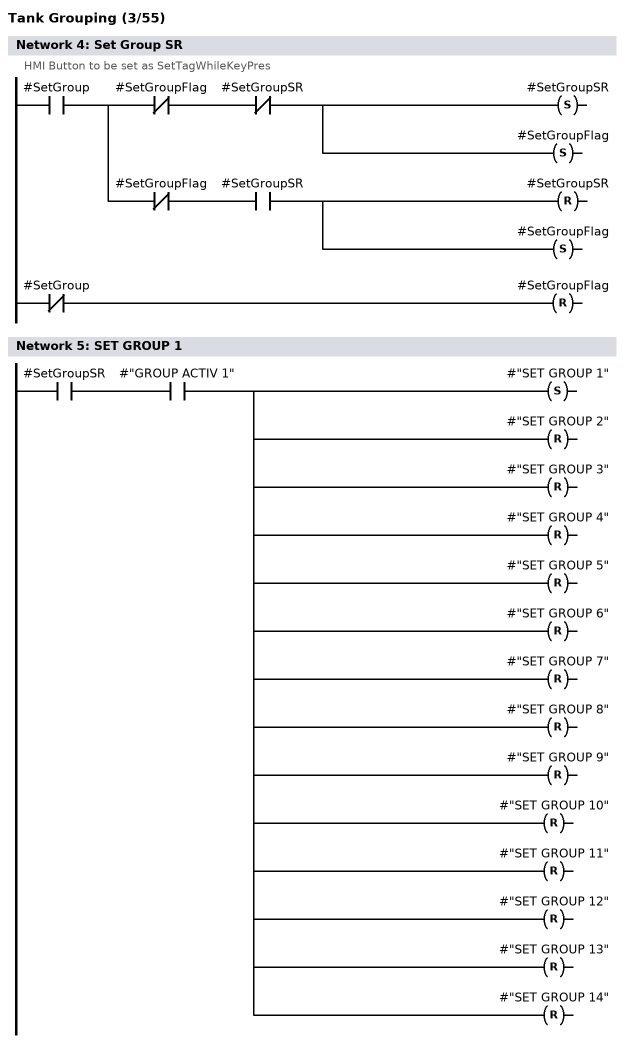
   RUNG wire#powerrail
      Contact( #SetGroup )
      wire#w1
      I_Contact( #SetGroupFlag )
      I_Contact( #SetGroupSR )
      wire#w2
      S_Coil( #SetGroupSR )
   END_RUNG
   RUNG wire#w2
      S_Coil( #SetGroupFlag )
   END_RUNG
   RUNG wire#w1
      I_Contact( #SetGroupFlag )
      Contact( #SetGroupSR )
      wire#w3
      R_Coil( #SetGroupSR )
   END_RUNG
   RUNG wire#w3
      S_Coil( #SetGroupFlag )
   END_RUNG
   RUNG wire#powerrail
      I_Contact( #SetGroup )
      R_Coil( #SetGroupFlag )
   END_RUNG
   // the same network as SCL:
   #_w1 := #SetGroup AND NOT #SetGroupFlag AND NOT #SetGroupSR;
   IF #_w1 THEN
       #SetGroupSR := TRUE;
       #SetGroupFlag := TRUE;
   END_IF;
   #_w2 := #SetGroup AND NOT #SetGroupFlag AND #SetGroupSR;
   IF #_w2 THEN
       #SetGroupSR := FALSE;
       #SetGroupFlag := TRUE;
   END_IF;
   IF NOT #SetGroup THEN #SetGroupFlag := FALSE; END_IF;
END_REGION

REGION Network 5: SET GROUP 1
   RUNG wire#powerrail
      Contact( #SetGroupSR )
      Contact( #"GROUP ACTIV 1" )
      wire#w1
      S_Coil( #"SET GROUP 1" )
   END_RUNG
   RUNG wire#w1
      R_Coil( #"SET GROUP 2" )
   END_RUNG
   RUNG wire#w1
      R_Coil( #"SET GROUP 3" )
   END_RUNG
   RUNG wire#w1
      R_Coil( #"SET GROUP 4" )
   END_RUNG
   RUNG wire#w1
      R_Coil( #"SET GROUP 5" )
   END_RUNG
   RUNG wire#w1
      R_Coil( #"SET GROUP 6" )
   END_RUNG
   RUNG wire#w1
      R_Coil( #"SET GROUP 7" )
   END_RUNG
   RUNG wire#w1
      R_Coil( #"SET GROUP 8" )
   END_RUNG
   RUNG wire#w1
      R_Coil( #"SET GROUP 9" )
   END_RUNG
   RUNG wire#w1
      R_Coil( #"SET GROUP 10" )
   END_RUNG
   RUNG wire#w1
      R_Coil( #"SET GROUP 11" )
   END_RUNG
   RUNG wire#w1
      R_Coil( #"SET GROUP 12" )
   END_RUNG
   RUNG wire#w1
      R_Coil( #"SET GROUP 13" )
   END_RUNG
   RUNG wire#w1
      R_Coil( #"SET GROUP 14" )
   END_RUNG
   // the same network as SCL:
   IF #SetGroupSR AND #"GROUP ACTIV 1" THEN
       #"SET GROUP 1" := TRUE;
       #"SET GROUP 2" := FALSE;
       #"SET GROUP 3" := FALSE;
       #"SET GROUP 4" := FALSE;
       #"SET GROUP 5" := FALSE;
       #"SET GROUP 6" := FALSE;
       #"SET GROUP 7" := FALSE;
       #"SET GROUP 8" := FALSE;
       #"SET GROUP 9" := FALSE;
       #"SET GROUP 10" := FALSE;
       #"SET GROUP 11" := FALSE;
       #"SET GROUP 12" := FALSE;
       #"SET GROUP 13" := FALSE;
       #"SET GROUP 14" := FALSE;
   END_IF;
END_REGION

REGION Network 6: SET GROUP 2
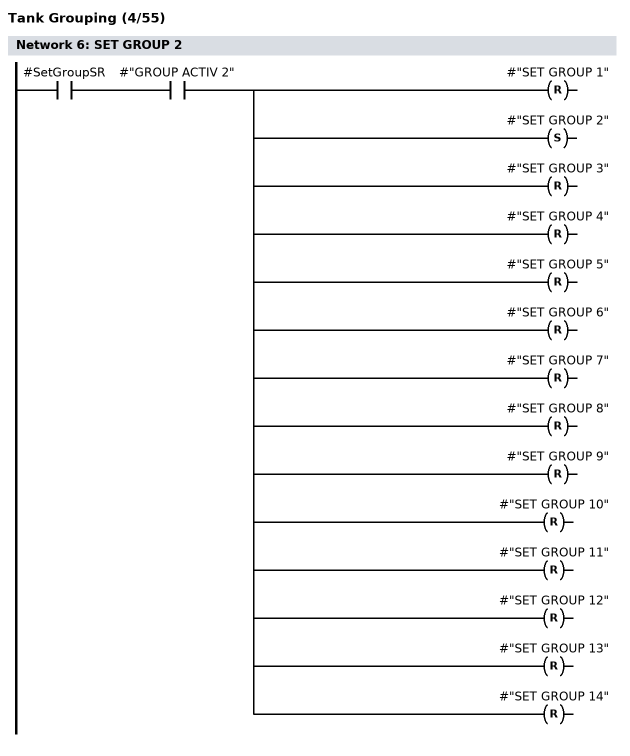
   RUNG wire#powerrail
      Contact( #SetGroupSR )
      Contact( #"GROUP ACTIV 2" )
      wire#w1
      R_Coil( #"SET GROUP 1" )
   END_RUNG
   RUNG wire#w1
      S_Coil( #"SET GROUP 2" )
   END_RUNG
   RUNG wire#w1
      R_Coil( #"SET GROUP 3" )
   END_RUNG
   RUNG wire#w1
      R_Coil( #"SET GROUP 4" )
   END_RUNG
   RUNG wire#w1
      R_Coil( #"SET GROUP 5" )
   END_RUNG
   RUNG wire#w1
      R_Coil( #"SET GROUP 6" )
   END_RUNG
   RUNG wire#w1
      R_Coil( #"SET GROUP 7" )
   END_RUNG
   RUNG wire#w1
      R_Coil( #"SET GROUP 8" )
   END_RUNG
   RUNG wire#w1
      R_Coil( #"SET GROUP 9" )
   END_RUNG
   RUNG wire#w1
      R_Coil( #"SET GROUP 10" )
   END_RUNG
   RUNG wire#w1
      R_Coil( #"SET GROUP 11" )
   END_RUNG
   RUNG wire#w1
      R_Coil( #"SET GROUP 12" )
   END_RUNG
   RUNG wire#w1
      R_Coil( #"SET GROUP 13" )
   END_RUNG
   RUNG wire#w1
      R_Coil( #"SET GROUP 14" )
   END_RUNG
   // the same network as SCL:
   IF #SetGroupSR AND #"GROUP ACTIV 2" THEN
       #"SET GROUP 1" := FALSE;
       #"SET GROUP 2" := TRUE;
       #"SET GROUP 3" := FALSE;
       #"SET GROUP 4" := FALSE;
       #"SET GROUP 5" := FALSE;
       #"SET GROUP 6" := FALSE;
       #"SET GROUP 7" := FALSE;
       #"SET GROUP 8" := FALSE;
       #"SET GROUP 9" := FALSE;
       #"SET GROUP 10" := FALSE;
       #"SET GROUP 11" := FALSE;
       #"SET GROUP 12" := FALSE;
       #"SET GROUP 13" := FALSE;
       #"SET GROUP 14" := FALSE;
   END_IF;
END_REGION

REGION Network 7: SET GROUP 3
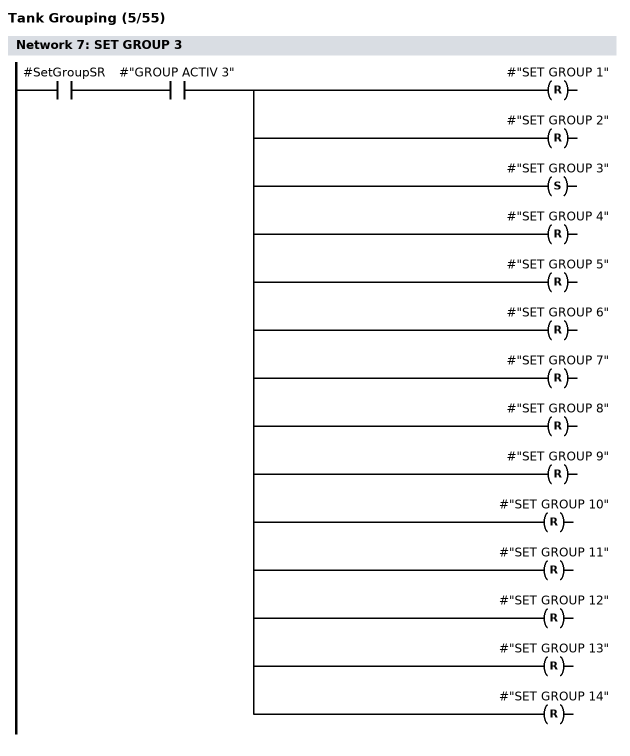
   RUNG wire#powerrail
      Contact( #SetGroupSR )
      Contact( #"GROUP ACTIV 3" )
      wire#w1
      R_Coil( #"SET GROUP 1" )
   END_RUNG
   RUNG wire#w1
      R_Coil( #"SET GROUP 2" )
   END_RUNG
   RUNG wire#w1
      S_Coil( #"SET GROUP 3" )
   END_RUNG
   RUNG wire#w1
      R_Coil( #"SET GROUP 4" )
   END_RUNG
   RUNG wire#w1
      R_Coil( #"SET GROUP 5" )
   END_RUNG
   RUNG wire#w1
      R_Coil( #"SET GROUP 6" )
   END_RUNG
   RUNG wire#w1
      R_Coil( #"SET GROUP 7" )
   END_RUNG
   RUNG wire#w1
      R_Coil( #"SET GROUP 8" )
   END_RUNG
   RUNG wire#w1
      R_Coil( #"SET GROUP 9" )
   END_RUNG
   RUNG wire#w1
      R_Coil( #"SET GROUP 10" )
   END_RUNG
   RUNG wire#w1
      R_Coil( #"SET GROUP 11" )
   END_RUNG
   RUNG wire#w1
      R_Coil( #"SET GROUP 12" )
   END_RUNG
   RUNG wire#w1
      R_Coil( #"SET GROUP 13" )
   END_RUNG
   RUNG wire#w1
      R_Coil( #"SET GROUP 14" )
   END_RUNG
   // the same network as SCL:
   IF #SetGroupSR AND #"GROUP ACTIV 3" THEN
       #"SET GROUP 1" := FALSE;
       #"SET GROUP 2" := FALSE;
       #"SET GROUP 3" := TRUE;
       #"SET GROUP 4" := FALSE;
       #"SET GROUP 5" := FALSE;
       #"SET GROUP 6" := FALSE;
       #"SET GROUP 7" := FALSE;
       #"SET GROUP 8" := FALSE;
       #"SET GROUP 9" := FALSE;
       #"SET GROUP 10" := FALSE;
       #"SET GROUP 11" := FALSE;
       #"SET GROUP 12" := FALSE;
       #"SET GROUP 13" := FALSE;
       #"SET GROUP 14" := FALSE;
   END_IF;
END_REGION

REGION Network 8: SET GROUP 4
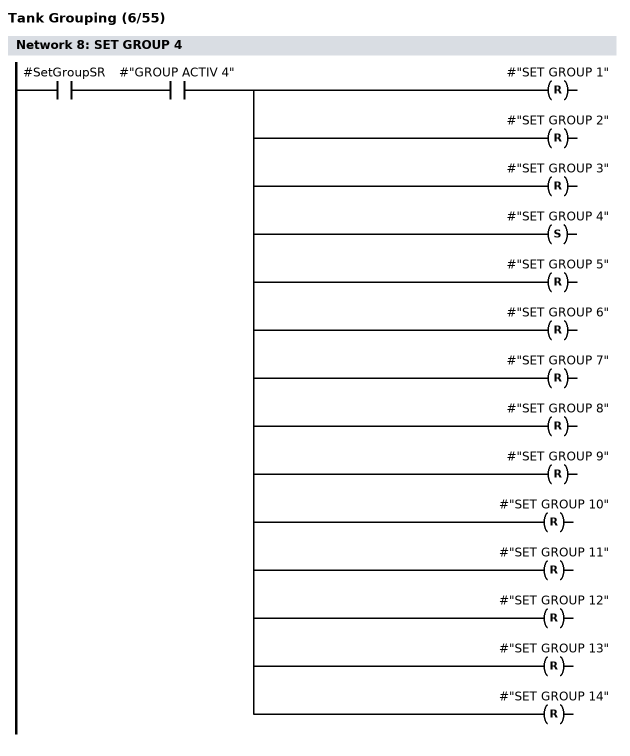
   RUNG wire#powerrail
      Contact( #SetGroupSR )
      Contact( #"GROUP ACTIV 4" )
      wire#w1
      R_Coil( #"SET GROUP 1" )
   END_RUNG
   RUNG wire#w1
      R_Coil( #"SET GROUP 2" )
   END_RUNG
   RUNG wire#w1
      R_Coil( #"SET GROUP 3" )
   END_RUNG
   RUNG wire#w1
      S_Coil( #"SET GROUP 4" )
   END_RUNG
   RUNG wire#w1
      R_Coil( #"SET GROUP 5" )
   END_RUNG
   RUNG wire#w1
      R_Coil( #"SET GROUP 6" )
   END_RUNG
   RUNG wire#w1
      R_Coil( #"SET GROUP 7" )
   END_RUNG
   RUNG wire#w1
      R_Coil( #"SET GROUP 8" )
   END_RUNG
   RUNG wire#w1
      R_Coil( #"SET GROUP 9" )
   END_RUNG
   RUNG wire#w1
      R_Coil( #"SET GROUP 10" )
   END_RUNG
   RUNG wire#w1
      R_Coil( #"SET GROUP 11" )
   END_RUNG
   RUNG wire#w1
      R_Coil( #"SET GROUP 12" )
   END_RUNG
   RUNG wire#w1
      R_Coil( #"SET GROUP 13" )
   END_RUNG
   RUNG wire#w1
      R_Coil( #"SET GROUP 14" )
   END_RUNG
   // the same network as SCL:
   IF #SetGroupSR AND #"GROUP ACTIV 4" THEN
       #"SET GROUP 1" := FALSE;
       #"SET GROUP 2" := FALSE;
       #"SET GROUP 3" := FALSE;
       #"SET GROUP 4" := TRUE;
       #"SET GROUP 5" := FALSE;
       #"SET GROUP 6" := FALSE;
       #"SET GROUP 7" := FALSE;
       #"SET GROUP 8" := FALSE;
       #"SET GROUP 9" := FALSE;
       #"SET GROUP 10" := FALSE;
       #"SET GROUP 11" := FALSE;
       #"SET GROUP 12" := FALSE;
       #"SET GROUP 13" := FALSE;
       #"SET GROUP 14" := FALSE;
   END_IF;
END_REGION

REGION Network 9: SET GROUP 5
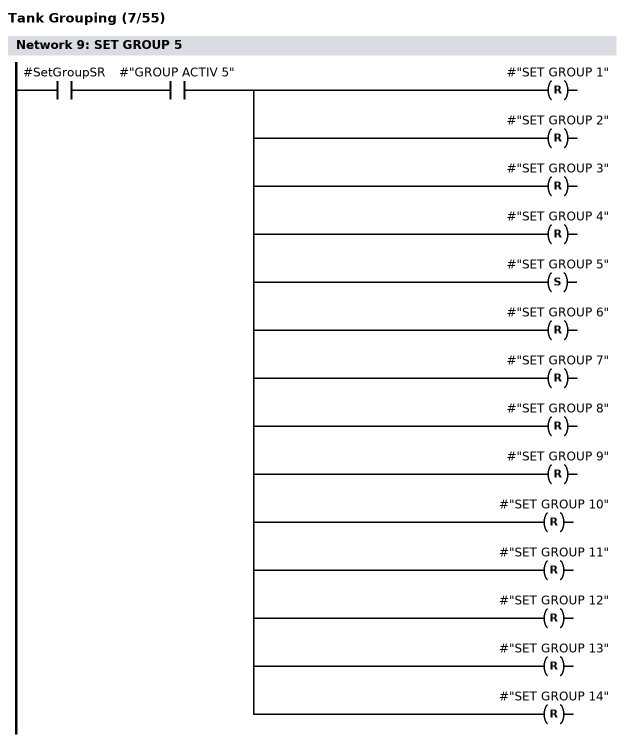
   RUNG wire#powerrail
      Contact( #SetGroupSR )
      Contact( #"GROUP ACTIV 5" )
      wire#w1
      R_Coil( #"SET GROUP 1" )
   END_RUNG
   RUNG wire#w1
      R_Coil( #"SET GROUP 2" )
   END_RUNG
   RUNG wire#w1
      R_Coil( #"SET GROUP 3" )
   END_RUNG
   RUNG wire#w1
      R_Coil( #"SET GROUP 4" )
   END_RUNG
   RUNG wire#w1
      S_Coil( #"SET GROUP 5" )
   END_RUNG
   RUNG wire#w1
      R_Coil( #"SET GROUP 6" )
   END_RUNG
   RUNG wire#w1
      R_Coil( #"SET GROUP 7" )
   END_RUNG
   RUNG wire#w1
      R_Coil( #"SET GROUP 8" )
   END_RUNG
   RUNG wire#w1
      R_Coil( #"SET GROUP 9" )
   END_RUNG
   RUNG wire#w1
      R_Coil( #"SET GROUP 10" )
   END_RUNG
   RUNG wire#w1
      R_Coil( #"SET GROUP 11" )
   END_RUNG
   RUNG wire#w1
      R_Coil( #"SET GROUP 12" )
   END_RUNG
   RUNG wire#w1
      R_Coil( #"SET GROUP 13" )
   END_RUNG
   RUNG wire#w1
      R_Coil( #"SET GROUP 14" )
   END_RUNG
   // the same network as SCL:
   IF #SetGroupSR AND #"GROUP ACTIV 5" THEN
       #"SET GROUP 1" := FALSE;
       #"SET GROUP 2" := FALSE;
       #"SET GROUP 3" := FALSE;
       #"SET GROUP 4" := FALSE;
       #"SET GROUP 5" := TRUE;
       #"SET GROUP 6" := FALSE;
       #"SET GROUP 7" := FALSE;
       #"SET GROUP 8" := FALSE;
       #"SET GROUP 9" := FALSE;
       #"SET GROUP 10" := FALSE;
       #"SET GROUP 11" := FALSE;
       #"SET GROUP 12" := FALSE;
       #"SET GROUP 13" := FALSE;
       #"SET GROUP 14" := FALSE;
   END_IF;
END_REGION

REGION Network 10: SET GROUP 6
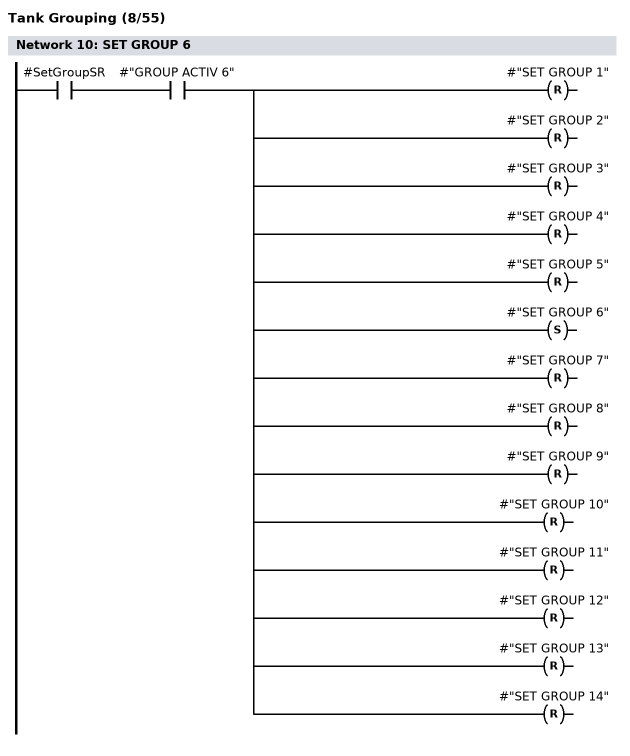
   RUNG wire#powerrail
      Contact( #SetGroupSR )
      Contact( #"GROUP ACTIV 6" )
      wire#w1
      R_Coil( #"SET GROUP 1" )
   END_RUNG
   RUNG wire#w1
      R_Coil( #"SET GROUP 2" )
   END_RUNG
   RUNG wire#w1
      R_Coil( #"SET GROUP 3" )
   END_RUNG
   RUNG wire#w1
      R_Coil( #"SET GROUP 4" )
   END_RUNG
   RUNG wire#w1
      R_Coil( #"SET GROUP 5" )
   END_RUNG
   RUNG wire#w1
      S_Coil( #"SET GROUP 6" )
   END_RUNG
   RUNG wire#w1
      R_Coil( #"SET GROUP 7" )
   END_RUNG
   RUNG wire#w1
      R_Coil( #"SET GROUP 8" )
   END_RUNG
   RUNG wire#w1
      R_Coil( #"SET GROUP 9" )
   END_RUNG
   RUNG wire#w1
      R_Coil( #"SET GROUP 10" )
   END_RUNG
   RUNG wire#w1
      R_Coil( #"SET GROUP 11" )
   END_RUNG
   RUNG wire#w1
      R_Coil( #"SET GROUP 12" )
   END_RUNG
   RUNG wire#w1
      R_Coil( #"SET GROUP 13" )
   END_RUNG
   RUNG wire#w1
      R_Coil( #"SET GROUP 14" )
   END_RUNG
   // the same network as SCL:
   IF #SetGroupSR AND #"GROUP ACTIV 6" THEN
       #"SET GROUP 1" := FALSE;
       #"SET GROUP 2" := FALSE;
       #"SET GROUP 3" := FALSE;
       #"SET GROUP 4" := FALSE;
       #"SET GROUP 5" := FALSE;
       #"SET GROUP 6" := TRUE;
       #"SET GROUP 7" := FALSE;
       #"SET GROUP 8" := FALSE;
       #"SET GROUP 9" := FALSE;
       #"SET GROUP 10" := FALSE;
       #"SET GROUP 11" := FALSE;
       #"SET GROUP 12" := FALSE;
       #"SET GROUP 13" := FALSE;
       #"SET GROUP 14" := FALSE;
   END_IF;
END_REGION

REGION Network 11: SET GROUP 7
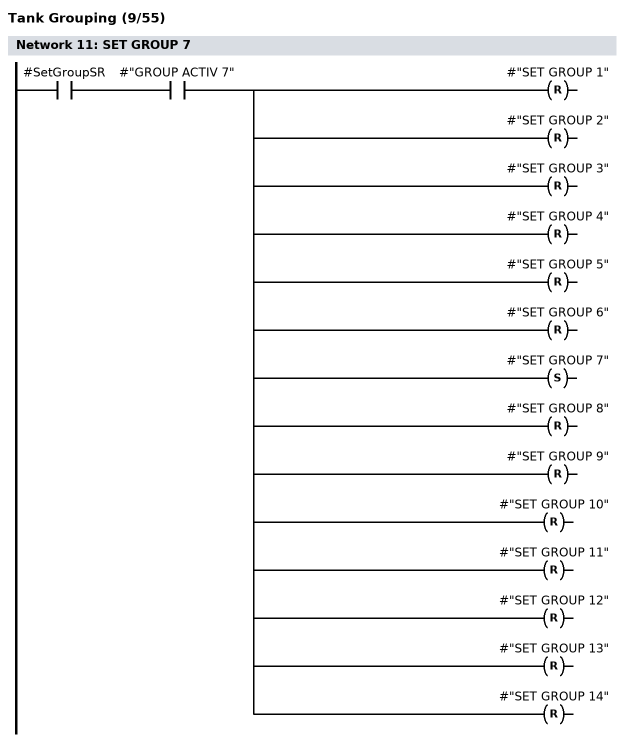
   RUNG wire#powerrail
      Contact( #SetGroupSR )
      Contact( #"GROUP ACTIV 7" )
      wire#w1
      R_Coil( #"SET GROUP 1" )
   END_RUNG
   RUNG wire#w1
      R_Coil( #"SET GROUP 2" )
   END_RUNG
   RUNG wire#w1
      R_Coil( #"SET GROUP 3" )
   END_RUNG
   RUNG wire#w1
      R_Coil( #"SET GROUP 4" )
   END_RUNG
   RUNG wire#w1
      R_Coil( #"SET GROUP 5" )
   END_RUNG
   RUNG wire#w1
      R_Coil( #"SET GROUP 6" )
   END_RUNG
   RUNG wire#w1
      S_Coil( #"SET GROUP 7" )
   END_RUNG
   RUNG wire#w1
      R_Coil( #"SET GROUP 8" )
   END_RUNG
   RUNG wire#w1
      R_Coil( #"SET GROUP 9" )
   END_RUNG
   RUNG wire#w1
      R_Coil( #"SET GROUP 10" )
   END_RUNG
   RUNG wire#w1
      R_Coil( #"SET GROUP 11" )
   END_RUNG
   RUNG wire#w1
      R_Coil( #"SET GROUP 12" )
   END_RUNG
   RUNG wire#w1
      R_Coil( #"SET GROUP 13" )
   END_RUNG
   RUNG wire#w1
      R_Coil( #"SET GROUP 14" )
   END_RUNG
   // the same network as SCL:
   IF #SetGroupSR AND #"GROUP ACTIV 7" THEN
       #"SET GROUP 1" := FALSE;
       #"SET GROUP 2" := FALSE;
       #"SET GROUP 3" := FALSE;
       #"SET GROUP 4" := FALSE;
       #"SET GROUP 5" := FALSE;
       #"SET GROUP 6" := FALSE;
       #"SET GROUP 7" := TRUE;
       #"SET GROUP 8" := FALSE;
       #"SET GROUP 9" := FALSE;
       #"SET GROUP 10" := FALSE;
       #"SET GROUP 11" := FALSE;
       #"SET GROUP 12" := FALSE;
       #"SET GROUP 13" := FALSE;
       #"SET GROUP 14" := FALSE;
   END_IF;
END_REGION

REGION Network 12: SET GROUP 8
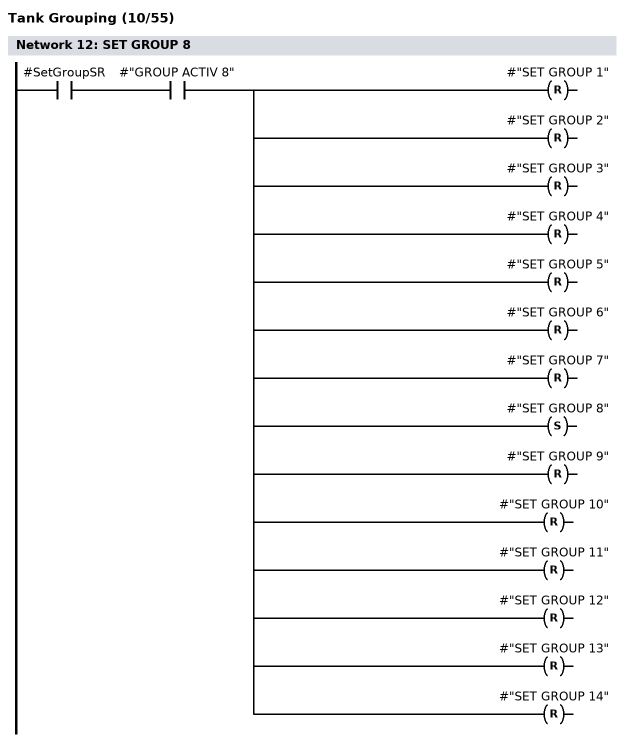
   RUNG wire#powerrail
      Contact( #SetGroupSR )
      Contact( #"GROUP ACTIV 8" )
      wire#w1
      R_Coil( #"SET GROUP 1" )
   END_RUNG
   RUNG wire#w1
      R_Coil( #"SET GROUP 2" )
   END_RUNG
   RUNG wire#w1
      R_Coil( #"SET GROUP 3" )
   END_RUNG
   RUNG wire#w1
      R_Coil( #"SET GROUP 4" )
   END_RUNG
   RUNG wire#w1
      R_Coil( #"SET GROUP 5" )
   END_RUNG
   RUNG wire#w1
      R_Coil( #"SET GROUP 6" )
   END_RUNG
   RUNG wire#w1
      R_Coil( #"SET GROUP 7" )
   END_RUNG
   RUNG wire#w1
      S_Coil( #"SET GROUP 8" )
   END_RUNG
   RUNG wire#w1
      R_Coil( #"SET GROUP 9" )
   END_RUNG
   RUNG wire#w1
      R_Coil( #"SET GROUP 10" )
   END_RUNG
   RUNG wire#w1
      R_Coil( #"SET GROUP 11" )
   END_RUNG
   RUNG wire#w1
      R_Coil( #"SET GROUP 12" )
   END_RUNG
   RUNG wire#w1
      R_Coil( #"SET GROUP 13" )
   END_RUNG
   RUNG wire#w1
      R_Coil( #"SET GROUP 14" )
   END_RUNG
   // the same network as SCL:
   IF #SetGroupSR AND #"GROUP ACTIV 8" THEN
       #"SET GROUP 1" := FALSE;
       #"SET GROUP 2" := FALSE;
       #"SET GROUP 3" := FALSE;
       #"SET GROUP 4" := FALSE;
       #"SET GROUP 5" := FALSE;
       #"SET GROUP 6" := FALSE;
       #"SET GROUP 7" := FALSE;
       #"SET GROUP 8" := TRUE;
       #"SET GROUP 9" := FALSE;
       #"SET GROUP 10" := FALSE;
       #"SET GROUP 11" := FALSE;
       #"SET GROUP 12" := FALSE;
       #"SET GROUP 13" := FALSE;
       #"SET GROUP 14" := FALSE;
   END_IF;
END_REGION

REGION Network 13: SET GROUP 9
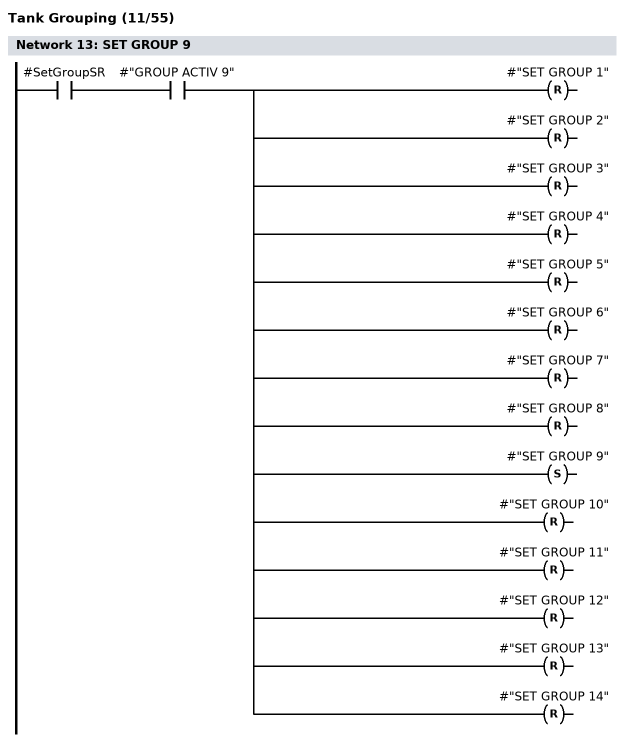
   RUNG wire#powerrail
      Contact( #SetGroupSR )
      Contact( #"GROUP ACTIV 9" )
      wire#w1
      R_Coil( #"SET GROUP 1" )
   END_RUNG
   RUNG wire#w1
      R_Coil( #"SET GROUP 2" )
   END_RUNG
   RUNG wire#w1
      R_Coil( #"SET GROUP 3" )
   END_RUNG
   RUNG wire#w1
      R_Coil( #"SET GROUP 4" )
   END_RUNG
   RUNG wire#w1
      R_Coil( #"SET GROUP 5" )
   END_RUNG
   RUNG wire#w1
      R_Coil( #"SET GROUP 6" )
   END_RUNG
   RUNG wire#w1
      R_Coil( #"SET GROUP 7" )
   END_RUNG
   RUNG wire#w1
      R_Coil( #"SET GROUP 8" )
   END_RUNG
   RUNG wire#w1
      S_Coil( #"SET GROUP 9" )
   END_RUNG
   RUNG wire#w1
      R_Coil( #"SET GROUP 10" )
   END_RUNG
   RUNG wire#w1
      R_Coil( #"SET GROUP 11" )
   END_RUNG
   RUNG wire#w1
      R_Coil( #"SET GROUP 12" )
   END_RUNG
   RUNG wire#w1
      R_Coil( #"SET GROUP 13" )
   END_RUNG
   RUNG wire#w1
      R_Coil( #"SET GROUP 14" )
   END_RUNG
   // the same network as SCL:
   IF #SetGroupSR AND #"GROUP ACTIV 9" THEN
       #"SET GROUP 1" := FALSE;
       #"SET GROUP 2" := FALSE;
       #"SET GROUP 3" := FALSE;
       #"SET GROUP 4" := FALSE;
       #"SET GROUP 5" := FALSE;
       #"SET GROUP 6" := FALSE;
       #"SET GROUP 7" := FALSE;
       #"SET GROUP 8" := FALSE;
       #"SET GROUP 9" := TRUE;
       #"SET GROUP 10" := FALSE;
       #"SET GROUP 11" := FALSE;
       #"SET GROUP 12" := FALSE;
       #"SET GROUP 13" := FALSE;
       #"SET GROUP 14" := FALSE;
   END_IF;
END_REGION

REGION Network 14: SET GROUP 10
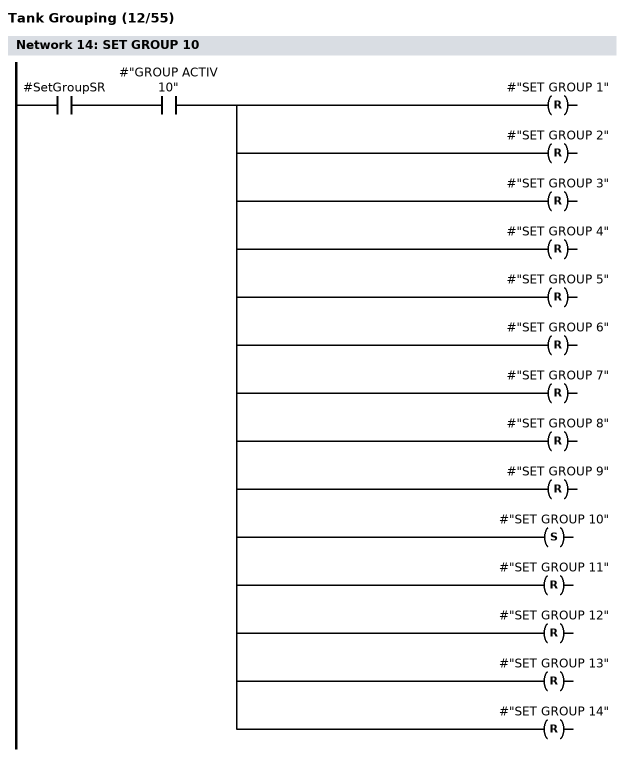
   RUNG wire#powerrail
      Contact( #SetGroupSR )
      Contact( #"GROUP ACTIV 10" )
      wire#w1
      R_Coil( #"SET GROUP 1" )
   END_RUNG
   RUNG wire#w1
      R_Coil( #"SET GROUP 2" )
   END_RUNG
   RUNG wire#w1
      R_Coil( #"SET GROUP 3" )
   END_RUNG
   RUNG wire#w1
      R_Coil( #"SET GROUP 4" )
   END_RUNG
   RUNG wire#w1
      R_Coil( #"SET GROUP 5" )
   END_RUNG
   RUNG wire#w1
      R_Coil( #"SET GROUP 6" )
   END_RUNG
   RUNG wire#w1
      R_Coil( #"SET GROUP 7" )
   END_RUNG
   RUNG wire#w1
      R_Coil( #"SET GROUP 8" )
   END_RUNG
   RUNG wire#w1
      R_Coil( #"SET GROUP 9" )
   END_RUNG
   RUNG wire#w1
      S_Coil( #"SET GROUP 10" )
   END_RUNG
   RUNG wire#w1
      R_Coil( #"SET GROUP 11" )
   END_RUNG
   RUNG wire#w1
      R_Coil( #"SET GROUP 12" )
   END_RUNG
   RUNG wire#w1
      R_Coil( #"SET GROUP 13" )
   END_RUNG
   RUNG wire#w1
      R_Coil( #"SET GROUP 14" )
   END_RUNG
   // the same network as SCL:
   IF #SetGroupSR AND #"GROUP ACTIV 10" THEN
       #"SET GROUP 1" := FALSE;
       #"SET GROUP 2" := FALSE;
       #"SET GROUP 3" := FALSE;
       #"SET GROUP 4" := FALSE;
       #"SET GROUP 5" := FALSE;
       #"SET GROUP 6" := FALSE;
       #"SET GROUP 7" := FALSE;
       #"SET GROUP 8" := FALSE;
       #"SET GROUP 9" := FALSE;
       #"SET GROUP 10" := TRUE;
       #"SET GROUP 11" := FALSE;
       #"SET GROUP 12" := FALSE;
       #"SET GROUP 13" := FALSE;
       #"SET GROUP 14" := FALSE;
   END_IF;
END_REGION

REGION Network 15: SET GROUP 11
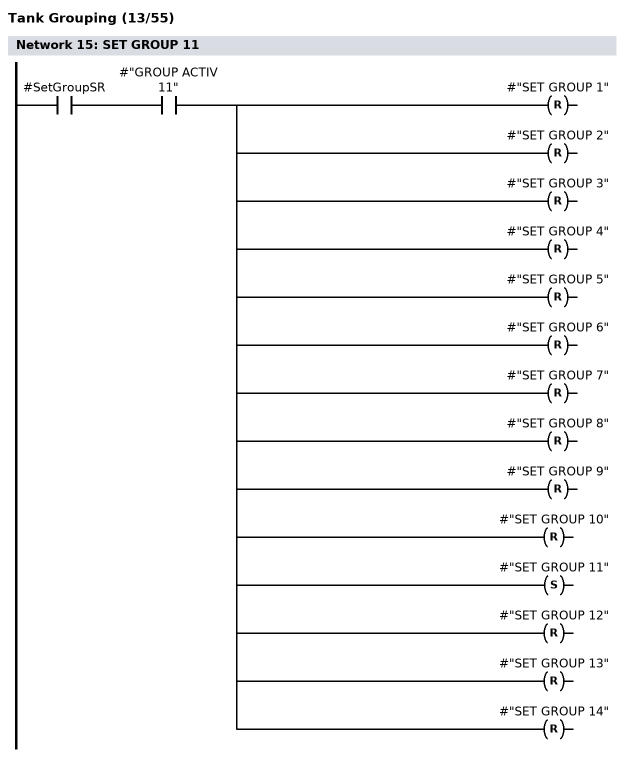
   RUNG wire#powerrail
      Contact( #SetGroupSR )
      Contact( #"GROUP ACTIV 11" )
      wire#w1
      R_Coil( #"SET GROUP 1" )
   END_RUNG
   RUNG wire#w1
      R_Coil( #"SET GROUP 2" )
   END_RUNG
   RUNG wire#w1
      R_Coil( #"SET GROUP 3" )
   END_RUNG
   RUNG wire#w1
      R_Coil( #"SET GROUP 4" )
   END_RUNG
   RUNG wire#w1
      R_Coil( #"SET GROUP 5" )
   END_RUNG
   RUNG wire#w1
      R_Coil( #"SET GROUP 6" )
   END_RUNG
   RUNG wire#w1
      R_Coil( #"SET GROUP 7" )
   END_RUNG
   RUNG wire#w1
      R_Coil( #"SET GROUP 8" )
   END_RUNG
   RUNG wire#w1
      R_Coil( #"SET GROUP 9" )
   END_RUNG
   RUNG wire#w1
      R_Coil( #"SET GROUP 10" )
   END_RUNG
   RUNG wire#w1
      S_Coil( #"SET GROUP 11" )
   END_RUNG
   RUNG wire#w1
      R_Coil( #"SET GROUP 12" )
   END_RUNG
   RUNG wire#w1
      R_Coil( #"SET GROUP 13" )
   END_RUNG
   RUNG wire#w1
      R_Coil( #"SET GROUP 14" )
   END_RUNG
   // the same network as SCL:
   IF #SetGroupSR AND #"GROUP ACTIV 11" THEN
       #"SET GROUP 1" := FALSE;
       #"SET GROUP 2" := FALSE;
       #"SET GROUP 3" := FALSE;
       #"SET GROUP 4" := FALSE;
       #"SET GROUP 5" := FALSE;
       #"SET GROUP 6" := FALSE;
       #"SET GROUP 7" := FALSE;
       #"SET GROUP 8" := FALSE;
       #"SET GROUP 9" := FALSE;
       #"SET GROUP 10" := FALSE;
       #"SET GROUP 11" := TRUE;
       #"SET GROUP 12" := FALSE;
       #"SET GROUP 13" := FALSE;
       #"SET GROUP 14" := FALSE;
   END_IF;
END_REGION

REGION Network 16: SET GROUP 12
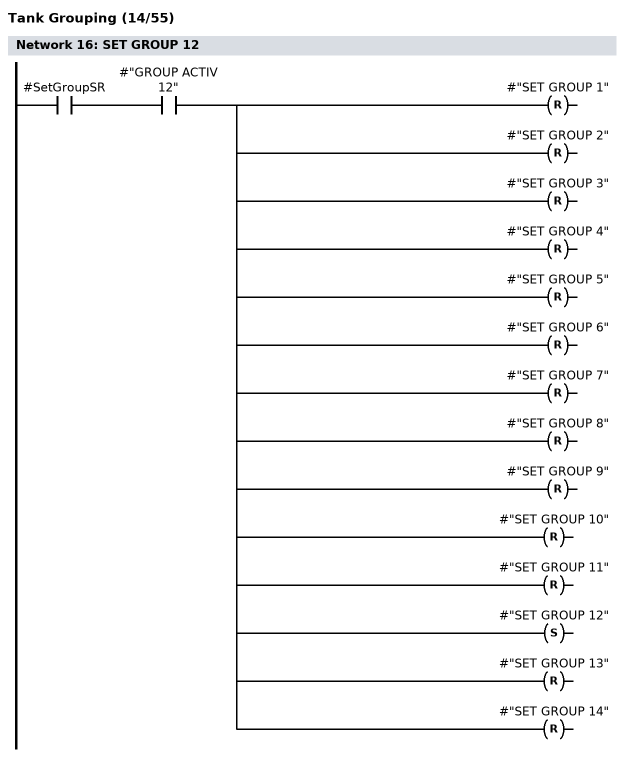
   RUNG wire#powerrail
      Contact( #SetGroupSR )
      Contact( #"GROUP ACTIV 12" )
      wire#w1
      R_Coil( #"SET GROUP 1" )
   END_RUNG
   RUNG wire#w1
      R_Coil( #"SET GROUP 2" )
   END_RUNG
   RUNG wire#w1
      R_Coil( #"SET GROUP 3" )
   END_RUNG
   RUNG wire#w1
      R_Coil( #"SET GROUP 4" )
   END_RUNG
   RUNG wire#w1
      R_Coil( #"SET GROUP 5" )
   END_RUNG
   RUNG wire#w1
      R_Coil( #"SET GROUP 6" )
   END_RUNG
   RUNG wire#w1
      R_Coil( #"SET GROUP 7" )
   END_RUNG
   RUNG wire#w1
      R_Coil( #"SET GROUP 8" )
   END_RUNG
   RUNG wire#w1
      R_Coil( #"SET GROUP 9" )
   END_RUNG
   RUNG wire#w1
      R_Coil( #"SET GROUP 10" )
   END_RUNG
   RUNG wire#w1
      R_Coil( #"SET GROUP 11" )
   END_RUNG
   RUNG wire#w1
      S_Coil( #"SET GROUP 12" )
   END_RUNG
   RUNG wire#w1
      R_Coil( #"SET GROUP 13" )
   END_RUNG
   RUNG wire#w1
      R_Coil( #"SET GROUP 14" )
   END_RUNG
   // the same network as SCL:
   IF #SetGroupSR AND #"GROUP ACTIV 12" THEN
       #"SET GROUP 1" := FALSE;
       #"SET GROUP 2" := FALSE;
       #"SET GROUP 3" := FALSE;
       #"SET GROUP 4" := FALSE;
       #"SET GROUP 5" := FALSE;
       #"SET GROUP 6" := FALSE;
       #"SET GROUP 7" := FALSE;
       #"SET GROUP 8" := FALSE;
       #"SET GROUP 9" := FALSE;
       #"SET GROUP 10" := FALSE;
       #"SET GROUP 11" := FALSE;
       #"SET GROUP 12" := TRUE;
       #"SET GROUP 13" := FALSE;
       #"SET GROUP 14" := FALSE;
   END_IF;
END_REGION

REGION Network 17: SET GROUP 13
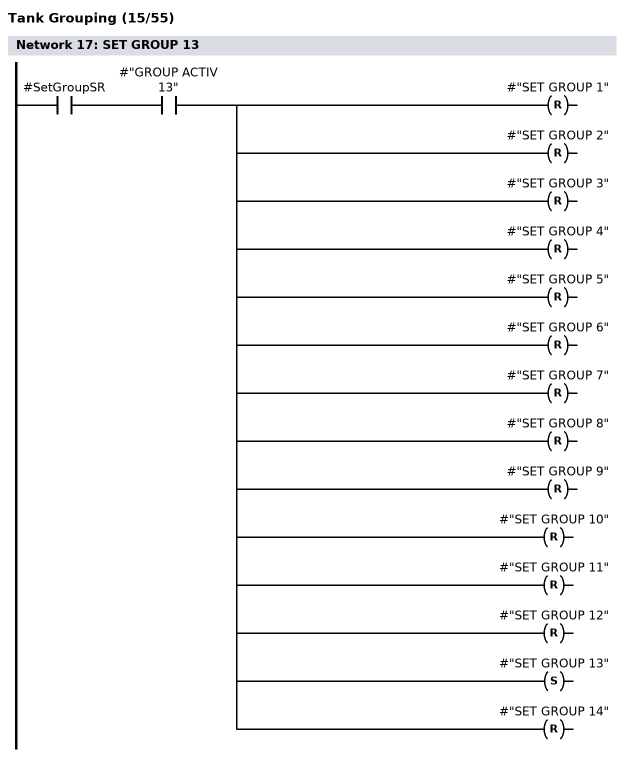
   RUNG wire#powerrail
      Contact( #SetGroupSR )
      Contact( #"GROUP ACTIV 13" )
      wire#w1
      R_Coil( #"SET GROUP 1" )
   END_RUNG
   RUNG wire#w1
      R_Coil( #"SET GROUP 2" )
   END_RUNG
   RUNG wire#w1
      R_Coil( #"SET GROUP 3" )
   END_RUNG
   RUNG wire#w1
      R_Coil( #"SET GROUP 4" )
   END_RUNG
   RUNG wire#w1
      R_Coil( #"SET GROUP 5" )
   END_RUNG
   RUNG wire#w1
      R_Coil( #"SET GROUP 6" )
   END_RUNG
   RUNG wire#w1
      R_Coil( #"SET GROUP 7" )
   END_RUNG
   RUNG wire#w1
      R_Coil( #"SET GROUP 8" )
   END_RUNG
   RUNG wire#w1
      R_Coil( #"SET GROUP 9" )
   END_RUNG
   RUNG wire#w1
      R_Coil( #"SET GROUP 10" )
   END_RUNG
   RUNG wire#w1
      R_Coil( #"SET GROUP 11" )
   END_RUNG
   RUNG wire#w1
      R_Coil( #"SET GROUP 12" )
   END_RUNG
   RUNG wire#w1
      S_Coil( #"SET GROUP 13" )
   END_RUNG
   RUNG wire#w1
      R_Coil( #"SET GROUP 14" )
   END_RUNG
   // the same network as SCL:
   IF #SetGroupSR AND #"GROUP ACTIV 13" THEN
       #"SET GROUP 1" := FALSE;
       #"SET GROUP 2" := FALSE;
       #"SET GROUP 3" := FALSE;
       #"SET GROUP 4" := FALSE;
       #"SET GROUP 5" := FALSE;
       #"SET GROUP 6" := FALSE;
       #"SET GROUP 7" := FALSE;
       #"SET GROUP 8" := FALSE;
       #"SET GROUP 9" := FALSE;
       #"SET GROUP 10" := FALSE;
       #"SET GROUP 11" := FALSE;
       #"SET GROUP 12" := FALSE;
       #"SET GROUP 13" := TRUE;
       #"SET GROUP 14" := FALSE;
   END_IF;
END_REGION

REGION Network 18: SET GROUP 14
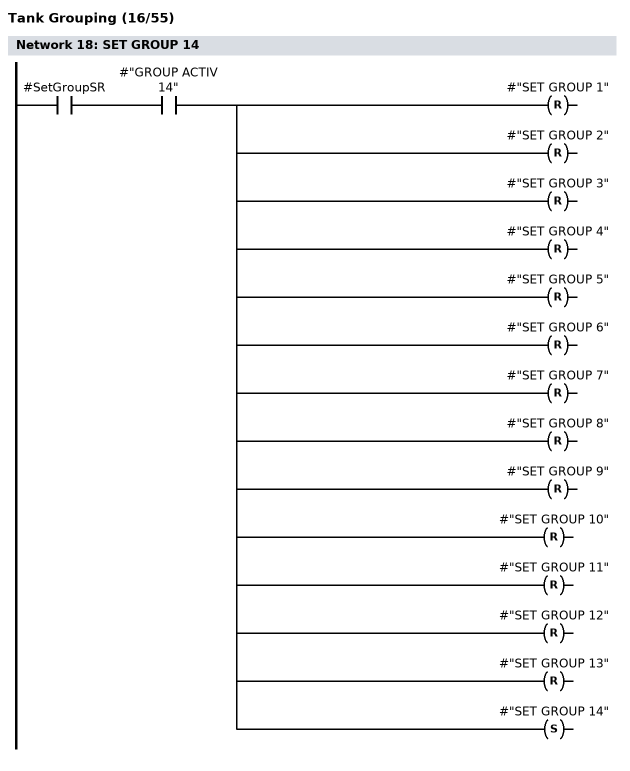
   RUNG wire#powerrail
      Contact( #SetGroupSR )
      Contact( #"GROUP ACTIV 14" )
      wire#w1
      R_Coil( #"SET GROUP 1" )
   END_RUNG
   RUNG wire#w1
      R_Coil( #"SET GROUP 2" )
   END_RUNG
   RUNG wire#w1
      R_Coil( #"SET GROUP 3" )
   END_RUNG
   RUNG wire#w1
      R_Coil( #"SET GROUP 4" )
   END_RUNG
   RUNG wire#w1
      R_Coil( #"SET GROUP 5" )
   END_RUNG
   RUNG wire#w1
      R_Coil( #"SET GROUP 6" )
   END_RUNG
   RUNG wire#w1
      R_Coil( #"SET GROUP 7" )
   END_RUNG
   RUNG wire#w1
      R_Coil( #"SET GROUP 8" )
   END_RUNG
   RUNG wire#w1
      R_Coil( #"SET GROUP 9" )
   END_RUNG
   RUNG wire#w1
      R_Coil( #"SET GROUP 10" )
   END_RUNG
   RUNG wire#w1
      R_Coil( #"SET GROUP 11" )
   END_RUNG
   RUNG wire#w1
      R_Coil( #"SET GROUP 12" )
   END_RUNG
   RUNG wire#w1
      R_Coil( #"SET GROUP 13" )
   END_RUNG
   RUNG wire#w1
      S_Coil( #"SET GROUP 14" )
   END_RUNG
   // the same network as SCL:
   IF #SetGroupSR AND #"GROUP ACTIV 14" THEN
       #"SET GROUP 1" := FALSE;
       #"SET GROUP 2" := FALSE;
       #"SET GROUP 3" := FALSE;
       #"SET GROUP 4" := FALSE;
       #"SET GROUP 5" := FALSE;
       #"SET GROUP 6" := FALSE;
       #"SET GROUP 7" := FALSE;
       #"SET GROUP 8" := FALSE;
       #"SET GROUP 9" := FALSE;
       #"SET GROUP 10" := FALSE;
       #"SET GROUP 11" := FALSE;
       #"SET GROUP 12" := FALSE;
       #"SET GROUP 13" := FALSE;
       #"SET GROUP 14" := TRUE;
   END_IF;
END_REGION

REGION Network 19: SET GROUP END
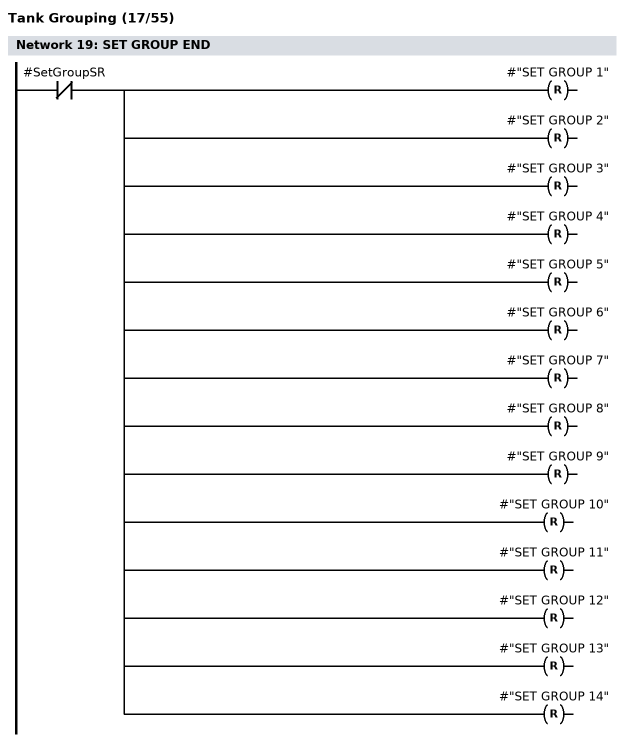
   RUNG wire#powerrail
      I_Contact( #SetGroupSR )
      wire#w1
      R_Coil( #"SET GROUP 1" )
   END_RUNG
   RUNG wire#w1
      R_Coil( #"SET GROUP 2" )
   END_RUNG
   RUNG wire#w1
      R_Coil( #"SET GROUP 3" )
   END_RUNG
   RUNG wire#w1
      R_Coil( #"SET GROUP 4" )
   END_RUNG
   RUNG wire#w1
      R_Coil( #"SET GROUP 5" )
   END_RUNG
   RUNG wire#w1
      R_Coil( #"SET GROUP 6" )
   END_RUNG
   RUNG wire#w1
      R_Coil( #"SET GROUP 7" )
   END_RUNG
   RUNG wire#w1
      R_Coil( #"SET GROUP 8" )
   END_RUNG
   RUNG wire#w1
      R_Coil( #"SET GROUP 9" )
   END_RUNG
   RUNG wire#w1
      R_Coil( #"SET GROUP 10" )
   END_RUNG
   RUNG wire#w1
      R_Coil( #"SET GROUP 11" )
   END_RUNG
   RUNG wire#w1
      R_Coil( #"SET GROUP 12" )
   END_RUNG
   RUNG wire#w1
      R_Coil( #"SET GROUP 13" )
   END_RUNG
   RUNG wire#w1
      R_Coil( #"SET GROUP 14" )
   END_RUNG
   // the same network as SCL:
   IF NOT #SetGroupSR THEN
       #"SET GROUP 1" := FALSE;
       #"SET GROUP 2" := FALSE;
       #"SET GROUP 3" := FALSE;
       #"SET GROUP 4" := FALSE;
       #"SET GROUP 5" := FALSE;
       #"SET GROUP 6" := FALSE;
       #"SET GROUP 7" := FALSE;
       #"SET GROUP 8" := FALSE;
       #"SET GROUP 9" := FALSE;
       #"SET GROUP 10" := FALSE;
       #"SET GROUP 11" := FALSE;
       #"SET GROUP 12" := FALSE;
       #"SET GROUP 13" := FALSE;
       #"SET GROUP 14" := FALSE;
   END_IF;
END_REGION

REGION Network 20: GROUP SET INDICATION